      Appearance <- "[78]"
   Button "Button_79" at 263,574 size 80x46; TextOff 'EMS 79'
      on Release: ActivateScreen("711_CARRIER_STATUS", 0)
      on Press: SetTag("HMI_EMS_Nr", 79)
      ObjectEnable <- "DB16_EMS_Status_EMS_DeviceStates.DeviceStates_Condition_HMI[79]"
      Appearance <- "[79]"
   Button "Button_80" at 346,574 size 80x46; TextOff 'EMS 80'
      on Release: ActivateScreen("711_CARRIER_STATUS", 0)
      on Press: SetTag("HMI_EMS_Nr", 80)
      ObjectEnable <- "DB16_EMS_Status_EMS_DeviceStates.DeviceStates_Condition_HMI[80]"
      Appearance <- "[80]"
   Button "Button_81" at 429,574 size 80x46; TextOff 'EMS 81'
      on Release: ActivateScreen("711_CARRIER_STATUS", 0)
      on Press: SetTag("HMI_EMS_Nr", 81)
      ObjectEnable <- "DB16_EMS_Status_EMS_DeviceStates.DeviceStates_Condition_HMI[81]"
      Appearance <- "[81]"
   Button "Button_82" at 512,574 size 80x46; TextOff 'EMS 82'
      on Release: ActivateScreen("711_CARRIER_STATUS", 0)
      on Press: SetTag("HMI_EMS_Nr", 82)
      ObjectEnable <- "DB16_EMS_Status_EMS_DeviceStates.DeviceStates_Condition_HMI[82]"
      Appearance <- "[82]"
   Button "Button_83" at 595,574 size 80x46; TextOff 'Text'
   Button "Button_84" at 678,574 size 80x46; TextOff 'Text'
   Button "Button_85" at 761,574 size 80x46; TextOff 'Text'
   Button "Button_86" at 845,574 size 80x46; TextOff 'Text'
   Button "Button_87" at 928,574 size 80x46; TextOff 'Text'
   Button "Button_88" at 1011,574 size 80x46; TextOff 'Text'
   Button "Button_89" at 1094,574 size 80x46; TextOff 'Text'
   Button "Button_90" at 1178,574 size 80x46; TextOff 'Text'
   TextField "Textfeld_7" at 567,118 size 243x27; Text 'section counter / min Barcode mm / EMS Status'
   TextField "Text field_1" at 83,642 size 97x25; Text 'NO COMM'
   TextField "Text field_2" at 83,683 size 191x25; Text 'ACTIVE, NO FAULTS'
   TextField "Text field_3" at 83,722 size 90x25; Text 'FAULTED'
   TextField "Text field_4" at 83,763 size 100x25; Text 'WARNING'

screen "700_System_Line_Overview" 1280x800
   GraphicView "Graphic view_1" at 0,119 size 1144x681; Picture "LAYOUT 1"
   TextField "Text field_126" at 847,138 size 285x28; Text 'SYSTEM LAYOUT SCREEN'
   Button "Template_Button_3" at 1074,2 size 203x55; TextOn 'FAULT RESET FAULT RESET'; TextOff 'FAULT RESET FAULT RESET'
      on Release: ResetBit("DB_SDC_GLOBAL_M.SDC_ER_Reset")
      on Press: SetBit("DB_SDC_GLOBAL_M.SDC_ER_Reset")
   AlarmView "Template_Alarm view_2" at 128,2 size 948x112
   Button "Template_Button_4" at 1196,56 size 81x59; TextOff 'Text'
      Appearance <- "AlwaysTRUE"
   Button "Button_21" at 0,57 size 128x58; TextOff 'SELECT SCREEN'
      on Release: ActivateScreen("010_START", 0)
   Button "Button_22" at 0,0 size 128x58; TextOff 'PREVIOUS SCREEN'
      on Click: function_efd93a16()
   DateTimeField "Template_Date/time field_2" at 1075,56 size 123x28
   DateTimeField "Template_Date/time field_3" at 1075,83 size 122x32
   TextField "Text field_2" at 446,600 size 186x29; Text 'Line Overview 1'
   TextField "Text field_3" at 524,179 size 186x29; Text 'Line Overview 3'
   TextField "Text field_4" at 564,383 size 186x29; Text 'Line Overview 2'
   TextField "Text field_5" at 811,383 size 186x29; Text 'Line Overview 4'
   Button "Button_1" at 436,216 size 134x49; TextOn 'LINE_OVERVIEW_2 LINE OVERVIEW_2'; TextOff 'LINE_OVERVIEW_2 LINE OVERVIEW_3'
      on Click: ActivateScreen("703_Line_Overview_3", 0)
   Button "Button_2" at 592,438 size 134x49; TextOn 'LINE_OVERVIEW_2 LINE OVERVIEW_2'; TextOff 'LINE_OVERVIEW_2 LINE OVERVIEW_2'
      on Click: ActivateScreen("702_Line_Overview_2", 0)
   Button "Button_3" at 840,438 size 134x49; TextOn 'LINE_OVERVIEW_2 LINE OVERVIEW_2'; TextOff 'LINE_OVERVIEW_2 LINE OVERVIEW_4'
      on Click: ActivateScreen("704_Line_Overview_4", 0)
   Button "Button_4" at 1148,702 size 127x87; TextOn 'LINE_OVERVIEW_2 LINE OVERVIEW_2'; TextOff 'LINE_OVERVIEW_2 / Main Screen'
      on Click: ActivateScreen("010_START", 0)
   Button "Button_14" at 247,578 size 134x49; TextOn 'LINE_OVERVIEW_2 LINE OVERVIEW_2'; TextOff 'LINE_OVERVIEW_2 LINE OVERVIEW_1'
      on Click: ActivateScreen("701_Line_Overview_1", 0)

screen "LINE_OVERVIEW_1_NOT_USED" 1280x800
   GraphicView "Graphic view_1" at 79,0 size 1139x766; Picture "b1 123927_1"
   TextField "Text field_1" at 981,284 size 46x25; Text 'S14'
   TextField "Text field_2" at 901,284 size 46x25; Text 'S13'
   TextField "Text field_3" at 818,283 size 46x25; Text 'S12'
   TextField "Text field_4" at 778,283 size 46x25; Text 'S11'
   TextField "Text field_5" at 734,283 size 46x25; Text 'S10'
   TextField "Text field_6" at 696,283 size 46x25; Text 'S9'
   TextField "Text field_7" at 653,283 size 46x25; Text 'S57'
   TextField "Text field_8" at 296,283 size 46x25; Text 'S7'
   TextField "Text field_9" at 252,283 size 46x25; Text 'S6'
   TextField "Text field_10" at 154,382 size 46x25; Text 'S5'
   TextField "Text field_11" at 245,471 size 46x25; Text 'S4'
   TextField "Text field_12" at 152,437 size 46x25; Text 'S3'
   TextField "Text field_13" at 22,532 size 46x25; Text 'S2'
   TextField "Text field_14" at 13,622 size 46x25; Text 'S58'
   TextField "Text field_15" at 22,671 size 46x25; Text 'S1'
   TextField "Text field_16" at 13,707 size 46x25; Text 'S56'
   TextField "Text field_17" at 128,721 size 46x25; Text 'S55'
   TextField "Text field_18" at 249,709 size 46x25; Text 'S54'
   TextField "Text field_19" at 212,590 size 46x25; Text 'S53'
   TextField "Text field_20" at 306,590 size 46x25; Text 'S52'
   TextField "Text field_21" at 395,591 size 46x25; Text 'S51'
   TextField "Text field_22" at 473,493 size 46x25; Text 'S47'
   TextField "Text field_23" at 544,492 size 46x25; Text 'S48'
   TextField "Text field_24" at 477,674 size 46x25; Text 'S44'
   TextField "Text field_25" at 546,674 size 46x25; Text 'S43'
   TextField "Text field_26" at 622,674 size 46x25; Text 'S42'
   TextField "Text field_27" at 723,641 size 46x25; Text 'S41'
   TextField "Text field_28" at 774,523 size 46x25; Text 'S40'
   TextField "Text field_29" at 883,607 size 46x25; Text 'S39'
   TextField "Text field_30" at 1015,607 size 46x25; Text 'S38'
   TextField "Text field_31" at 1114,607 size 46x25; Text 'S37'
   TextField "Text field_32" at 1158,502 size 46x25; Text 'S36'
   TextField "Text field_33" at 1157,438 size 46x25; Text 'S35'
   TextField "Text field_34" at 1158,381 size 46x25; Text 'S34'
   TextField "Text field_35" at 33,44 size 84x24; Text 'Area Name'
   TextField "Text field_36" at 36,62 size 56x25; Text 'Area A'
   Button "Button_14" at 980,678 size 140x105; TextOn 'LINE_OVERVIEW_2 LINE OVERVIEW_2'; TextOff 'LINE_OVERVIEW_2 LINE OVERVIEW_2'
      on Click: ActivateScreen("LINE_OVERVIEW_2_NOT_USED", 0)
   Button "Button_1" at 1125,677 size 140x105; TextOn 'LINE_OVERVIEW_2 LINE OVERVIEW_2'; TextOff 'LINE_OVERVIEW_2 / Main Screen'
      on Click: ActivateScreen("010_START", 0)
   TextField "Text field_37" at 36,78 size 67x25; Text 'Area AA'
   TextField "Text field_38" at 36,94 size 55x25; Text 'Area B'
   TextField "Text field_39" at 36,112 size 65x25; Text 'Area BB'
   TextField "Text field_40" at 36,129 size 55x25; Text 'Area C'
   TextField "Text field_41" at 36,147 size 65x25; Text 'Area CC'
   TextField "Text field_42" at 36,165 size 56x25; Text 'Area H'
   TextField "Text field_43" at 36,182 size 57x25; Text 'Area D'
   TextField "Text field_44" at 36,200 size 55x25; Text 'Area E'
   TextField "Text field_45" at 36,218 size 54x25; Text 'Area F'
   TextField "Text field_46" at 36,237 size 63x25; Text 'Area FF'
   TextField "Text field_47" at 36,256 size 56x25; Text 'Area G'
   TextField "Text field_48" at 242,42 size 81x26; Text 'Area Start'
   TextField "Text field_49" at 241,61 size 109x25; Text 'After Cab Pick'
   TextField "Text field_50" at 241,77 size 39x25; Text 'DL 1'
   TextField "Text field_51" at 241,94 size 155x25; Text 'DL 2 (Marriege Cell)'
   TextField "Text field_52" at 240,111 size 166x25; Text 'S14 at 90 degree turn'
   TextField "Text field_53" at 240,128 size 123x25; Text 'S16 Check Point'
   TextField "Text field_54" at 240,147 size 187x25; Text 'S19 above Front Bumper'
   TextField "Text field_55" at 240,164 size 125x25; Text 'from the Shuttle'
   TextField "Text field_56" at 240,181 size 169x25; Text 'S32 at 90 Degree turn'
   TextField "Text field_57" at 240,200 size 192x25; Text 'S33 at EMS01 Main Panel'
   TextField "Text field_58" at 240,219 size 198x25; Text 'S36 before 90 degree turn'
   TextField "Text field_59" at 241,237 size 106x25; Text 'Before Repair'
   TextField "Text field_60" at 241,255 size 91x25; Text 'Repair Spur'
   TextField "Text field_61" at 445,43 size 73x26; Text 'Area End'
   TextField "Text field_62" at 445,62 size 38x25; Text 'DL1'
   TextField "Text field_63" at 445,77 size 155x25; Text 'DL 2 (Marriege Cell)'
   TextField "Text field_64" at 445,95 size 166x25; Text 'S14 at 90 degree turn'
   TextField "Text field_65" at 445,113 size 123x25; Text 'S16 Check Point'
   TextField "Text field_66" at 445,130 size 187x25; Text 'S19 above Front Bumper'
   TextField "Text field_67" at 445,147 size 139x25; Text 'Before the Shuttle'
   TextField "Text field_68" at 444,165 size 169x25; Text 'S32 at 90 Degree turn'
   TextField "Text field_69" at 444,183 size 192x25; Text 'S33 at EMS01 Main Panel'
   TextField "Text field_70" at 444,201 size 198x25; Text 'S36 before 90 degree turn'
   TextField "Text field_71" at 445,220 size 106x25; Text 'Before Repair'
   TextField "Text field_72" at 446,238 size 67x25; Text 'Cab Pick'
   TextField "Text field_73" at 446,255 size 91x25; Text 'Repair Spur'
   TextField "Text field_74" at 652,43 size 67x26; Text 'Location'
   TextField "Text field_75" at 651,62 size 45x25; Text '@G7'
   TextField "Text field_76" at 651,79 size 47x25; Text '@F14'
   TextField "Text field_77" at 651,96 size 47x25; Text '@F14'
   TextField "Text field_78" at 651,112 size 50x25; Text '@Q16'
   TextField "Text field_79" at 651,131 size 50x25; Text '@Q16'
   TextField "Text field_80" at 651,149 size 49x25; Text '@U12'
   TextField "Text field_81" at 651,167 size 49x25; Text '@U12'
   TextField "Text field_82" at 651,184 size 46x25; Text '@L17'
   TextField "Text field_83" at 651,202 size 46x25; Text '@L17'
   TextField "Text field_84" at 651,221 size 48x25; Text '@C17'
   TextField "Text field_85" at 651,239 size 41x25; Text '@D9'
   TextField "Text field_86" at 651,257 size 41x25; Text '@D9'
   TextField "Text field_87" at 737,42 size 45x26; Text 'Panel'
   TextField "Text field_88" at 736,62 size 115x25; Text 'EMS01R2 JB33'
   TextField "Text field_89" at 736,80 size 75x25; Text 'EMS01R3'
   TextField "Text field_90" at 736,97 size 75x25; Text 'EMS01R3'
   TextField "Text field_91" at 736,113 size 100x25; Text 'EMS01 JB22'
   TextField "Text field_92" at 736,130 size 95x25; Text 'EMS01 JB22'
   TextField "Text field_93" at 736,148 size 75x25; Text 'EMS01R4'
   TextField "Text field_94" at 736,167 size 75x25; Text 'EMS01R4'
   TextField "Text field_95" at 736,185 size 55x25; Text 'EMS01'
   TextField "Text field_96" at 737,202 size 55x25; Text 'EMS01'
   TextField "Text field_97" at 737,220 size 115x25; Text 'EMS01R1 JB23'
   TextField "Text field_98" at 737,238 size 75x25; Text 'EMS01R1'
   TextField "Text field_99" at 737,256 size 75x25; Text 'EMS01R1'
   TextField "Text field_100" at 906,43 size 50x26; Text 'Offset'
   TextField "Text field_101" at 907,62 size 38x25; Text '9'
   TextField "Text field_102" at 907,80 size 38x25; Text '1'
   TextField "Text field_103" at 907,98 size 38x25; Text '2'
   TextField "Text field_104" at 907,114 size 38x25; Text '10'
   TextField "Text field_105" at 907,130 size 38x25; Text '11'
   TextField "Text field_106" at 907,150 size 38x25; Text '3'
   TextField "Text field_107" at 907,168 size 38x25; Text '4'
   TextField "Text field_108" at 907,185 size 38x25; Text '5'
   TextField "Text field_109" at 907,202 size 38x25; Text '6'
   TextField "Text field_110" at 907,221 size 38x25; Text '7'
   TextField "Text field_111" at 908,238 size 38x25; Text '12'
   TextField "Text field_112" at 908,256 size 38x25; Text '8'
   TextField "Text field_113" at 1084,54 size 82x22; Text 'AREA BB'
   TextField "Text field_114" at 1131,251 size 71x22; Text 'AREA E'
   TextField "Text field_115" at 940,613 size 71x22; Text 'AREA F'
   TextField "Text field_116" at 493,464 size 71x22; Text 'AREA G'
   TextField "Text field_117" at 267,679 size 82x22; Text 'AREA FF'
   TextField "Text field_118" at 138,519 size 71x22; Text 'AREA A'
   TextField "Text field_119" at 515,360 size 82x22; Text 'AREA AA'
   TextField "Text field_120" at 950,362 size 71x22; Text 'AREA B'
   TextField "Text field_121" at 731,358 size 53x27; Text 'DL2'
   TextField "Text field_122" at 712,381 size 93x25; Text 'Mrg Cell'
   TextField "Text field_123" at 296,359 size 53x27; Text 'DL1'
   TextField "Text field_124" at 125,635 size 49x25; Text 'Cab'
   TextField "Text field_125" at 125,656 size 49x25; Text 'Pick'
   TextField "Text field_126" at 454,13 size 341x28; Text 'OVERVIEW 1 - SCREEN 0023'
   TextField "Text field_127" at 614,387 size 82x24; Text 'EMS01R3'
   TextField "Text field_128" at 614,421 size 82x22; Text 'AREA AA'
   TextField "Text field_129" at 619,452 size 71x22; Text 'AREA B'
   TextField "Text field_130" at 23,313 size 82x24; Text 'EMS01R2'
   TextField "Text field_131" at 38,329 size 49x24; Text 'JB33'
   TextField "Text field_132" at 28,361 size 71x22; Text 'AREA A'
   TextField "Text field_133" at 379,679 size 82x24; Text 'EMS01R1'
   TextField "Text field_134" at 385,702 size 71x22; Text 'AREA G'
   TextField "Text field_135" at 386,729 size 71x22; Text 'AREA F'
   TextField "Text field_136" at 380,754 size 82x22; Text 'AREA FF'
   TextField "Text field_137" at 703,687 size 60x24; Text 'EMS01'
   TextField "Text field_138" at 699,718 size 71x22; Text 'AREA D'
   TextField "Text field_139" at 699,746 size 71x22; Text 'AREA E'
   TextField "Text field_140" at 790,686 size 82x24; Text 'EMS01R4'
   TextField "Text field_143" at 897,679 size 60x24; Text 'EMS01'
   TextField "Text field_144" at 902,693 size 49x24; Text 'JB22'
   DateTimeField "Date/time field_1" at 11,12 size 258x34
   TextField "Text field_141" at 790,718 size 82x22; Text 'AREA CC'
   TextField "Text field_142" at 796,746 size 71x22; Text 'AREA H'
   TextField "Text field_146" at 891,745 size 71x22; Text 'AREA C'
   TextField "Text field_145" at 886,718 size 82x22; Text 'AREA BB'
   TextField "Text field_147" at 863,43 size 38x26; Text 'Slot'
   TextField "Text field_148" at 865,62 size 38x25; Text '13'
   TextField "Text field_149" at 865,80 size 38x25; Text '5'
   TextField "Text field_150" at 865,97 size 38x25; Text '6'
   TextField "Text field_151" at 865,113 size 38x25; Text '14'
   TextField "Text field_152" at 865,131 size 38x25; Text '15'
   TextField "Text field_153" at 865,150 size 38x25; Text '7'
   TextField "Text field_154" at 865,166 size 38x25; Text '12'
   TextField "Text field_155" at 865,184 size 38x25; Text '8'
   TextField "Text field_156" at 865,202 size 38x25; Text '9'
   TextField "Text field_157" at 865,220 size 38x25; Text '10'
   TextField "Text field_158" at 866,238 size 38x25; Text '16'
   TextField "Text field_159" at 866,256 size 38x25; Text '11'
   TextField "Text field_160" at 120,43 size 40x26; Text 'Area'
   TextField "Text field_161" at 118,62 size 98x25; Text 'Cab Delivery'
   TextField "Text field_162" at 118,78 size 53x25; Text 'Trim 5'
   TextField "Text field_163" at 118,93 size 106x25; Text 'Body Delivery'
   TextField "Text field_164" at 118,110 size 106x25; Text 'Body Delivery'
   TextField "Text field_165" at 118,127 size 106x25; Text 'Body Delivery'
   TextField "Text field_166" at 118,146 size 106x25; Text 'Body Delivery'
   TextField "Text field_167" at 118,164 size 83x25; Text 'Body Deck'
   TextField "Text field_168" at 118,181 size 107x25; Text 'Empty Return'
   TextField "Text field_169" at 118,200 size 107x25; Text 'Empty Return'
   TextField "Text field_170" at 118,218 size 107x25; Text 'Empty Return'
   TextField "Text field_171" at 118,236 size 107x25; Text 'Empty Return'
   TextField "Text field_172" at 116,255 size 91x25; Text 'Repair Spur'
   IOField "I/O field_42" at 129,761 size 37x32; FormatPattern 99
      ProcessValue <- "CarrierNumber"
   IOField "I/O field_1" at 56,703 size 37x32; FormatPattern 99
      ProcessValue <- "CarrierNumber"
   IOField "I/O field_2" at 56,666 size 37x32; FormatPattern 99
      ProcessValue <- "CarrierNumber"
   IOField "I/O field_3" at 56,617 size 37x32; FormatPattern 99
      ProcessValue <- "CarrierNumber"
   IOField "I/O field_4" at 56,568 size 37x32; FormatPattern 99
      ProcessValue <- "CarrierNumber"
   IOField "I/O field_5" at 56,527 size 37x32; FormatPattern 99
      ProcessValue <- "CarrierNumber"
   IOField "I/O field_6" at 106,467 size 37x32; FormatPattern 99
      ProcessValue <- "CarrierNumber"
   IOField "I/O field_7" at 148,467 size 37x32; FormatPattern 99
      ProcessValue <- "CarrierNumber"
   IOField "I/O field_8" at 190,467 size 37x32; FormatPattern 99
      ProcessValue <- "CarrierNumber"
   IOField "I/O field_9" at 191,413 size 37x32; FormatPattern 99
      ProcessValue <- "CarrierNumber"
   IOField "I/O field_10" at 191,378 size 37x32; FormatPattern 99
      ProcessValue <- "CarrierNumber"
   IOField "I/O field_11" at 248,310 size 37x32; FormatPattern 99
      ProcessValue <- "CarrierNumber"
   IOField "I/O field_12" at 292,310 size 37x32; FormatPattern 99
      ProcessValue <- "CarrierNumber"
   IOField "I/O field_13" at 337,310 size 37x32; FormatPattern 99
      ProcessValue <- "CarrierNumber"
   IOField "I/O field_14" at 376,310 size 37x32; FormatPattern 99
      ProcessValue <- "CarrierNumber"
   IOField "I/O field_15" at 415,310 size 37x32; FormatPattern 99
      ProcessValue <- "CarrierNumber"
   IOField "I/O field_16" at 453,310 size 37x32; FormatPattern 99
      ProcessValue <- "CarrierNumber"
   IOField "I/O field_17" at 492,310 size 37x32; FormatPattern 99
      ProcessValue <- "CarrierNumber"
   IOField "I/O field_18" at 531,310 size 37x32; FormatPattern 99
      ProcessValue <- "CarrierNumber"
   IOField "I/O field_19" at 570,310 size 37x32; FormatPattern 99
      ProcessValue <- "CarrierNumber"
   IOField "I/O field_20" at 609,310 size 37x32; FormatPattern 99
      ProcessValue <- "CarrierNumber"
   IOField "I/O field_21" at 654,310 size 37x32; FormatPattern 99
      ProcessValue <- "CarrierNumber"
   IOField "I/O field_22" at 692,310 size 37x32; FormatPattern 99
      ProcessValue <- "CarrierNumber"
   IOField "I/O field_23" at 736,310 size 37x32; FormatPattern 99
      ProcessValue <- "CarrierNumber"
   IOField "I/O field_24" at 778,310 size 37x32; FormatPattern 99
      ProcessValue <- "CarrierNumber"
   IOField "I/O field_25" at 819,310 size 37x32; FormatPattern 99
      ProcessValue <- "CarrierNumber"
   IOField "I/O field_26" at 863,310 size 37x32; FormatPattern 99
      ProcessValue <- "CarrierNumber"
   IOField "I/O field_27" at 902,310 size 37x32; FormatPattern 99
      ProcessValue <- "CarrierNumber"
   IOField "I/O field_28" at 945,310 size 37x32; FormatPattern 99
      ProcessValue <- "CarrierNumber"
   IOField "I/O field_29" at 984,310 size 37x32; FormatPattern 99
      ProcessValue <- "CarrierNumber"
   IOField "I/O field_30" at 1031,289 size 37x32; FormatPattern 99
      ProcessValue <- "CarrierNumber"
   IOField "I/O field_31" at 1031,257 size 37x32; FormatPattern 99
      ProcessValue <- "CarrierNumber"
   IOField "I/O field_32" at 1031,225 size 37x32; FormatPattern 99
      ProcessValue <- "CarrierNumber"
   IOField "I/O field_33" at 1031,193 size 37x32; FormatPattern 99
      ProcessValue <- "CarrierNumber"
   IOField "I/O field_34" at 1031,162 size 37x32; FormatPattern 99
      ProcessValue <- "CarrierNumber"
   IOField "I/O field_35" at 1031,131 size 37x32; FormatPattern 99
      ProcessValue <- "CarrierNumber"
   IOField "I/O field_36" at 1031,99 size 37x32; FormatPattern 99
      ProcessValue <- "CarrierNumber"
   IOField "I/O field_37" at 1031,67 size 37x32; FormatPattern 99
      ProcessValue <- "CarrierNumber"
   IOField "I/O field_38" at 1031,35 size 37x32; FormatPattern 99
      ProcessValue <- "CarrierNumber"
   IOField "I/O field_39" at 1031,3 size 37x32; FormatPattern 99
      ProcessValue <- "CarrierNumber"
   IOField "I/O field_49" at 1219,339 size 37x32; FormatPattern 99
      ProcessValue <- "CarrierNumber"
   IOField "I/O field_50" at 1219,378 size 37x32; FormatPattern 99
      ProcessValue <- "CarrierNumber"
   IOField "I/O field_51" at 1219,435 size 37x32; FormatPattern 99
      ProcessValue <- "CarrierNumber"
   IOField "I/O field_52" at 1218,498 size 37x32; FormatPattern 99
      ProcessValue <- "CarrierNumber"
   IOField "I/O field_40" at 1218,302 size 37x32; FormatPattern 99
      ProcessValue <- "CarrierNumber"
   IOField "I/O field_41" at 1218,265 size 37x32; FormatPattern 99
      ProcessValue <- "CarrierNumber"
   IOField "I/O field_43" at 1218,228 size 37x32; FormatPattern 99
      ProcessValue <- "CarrierNumber"
   IOField "I/O field_44" at 1218,191 size 37x32; FormatPattern 99
      ProcessValue <- "CarrierNumber"
   IOField "I/O field_45" at 1218,154 size 37x32; FormatPattern 99
      ProcessValue <- "CarrierNumber"
   IOField "I/O field_46" at 1218,117 size 37x32; FormatPattern 99
      ProcessValue <- "CarrierNumber"
   IOField "I/O field_47" at 1218,80 size 37x32; FormatPattern 99
      ProcessValue <- "CarrierNumber"
   IOField "I/O field_48" at 1218,43 size 37x32; FormatPattern 99
      ProcessValue <- "CarrierNumber"
   IOField "I/O field_53" at 1156,568 size 37x32; FormatPattern 99
      ProcessValue <- "CarrierNumber"
   IOField "I/O field_54" at 1115,568 size 37x32; FormatPattern 99
      ProcessValue <- "CarrierNumber"
   IOField "I/O field_55" at 1054,568 size 37x32; FormatPattern 99
      ProcessValue <- "CarrierNumber"
   IOField "I/O field_56" at 1015,568 size 37x32; FormatPattern 99
      ProcessValue <- "CarrierNumber"
   IOField "I/O field_57" at 924,568 size 37x32; FormatPattern 99
      ProcessValue <- "CarrierNumber"
   IOField "I/O field_58" at 884,568 size 37x32; FormatPattern 99
      ProcessValue <- "CarrierNumber"
   IOField "I/O field_59" at 813,568 size 37x32; FormatPattern 99
      ProcessValue <- "CarrierNumber"
   IOField "I/O field_60" at 773,568 size 37x32; FormatPattern 99
      ProcessValue <- "CarrierNumber"
   IOField "I/O field_61" at 724,603 size 37x32; FormatPattern 99
      ProcessValue <- "CarrierNumber"
   IOField "I/O field_62" at 663,634 size 37x32; FormatPattern 99
      ProcessValue <- "CarrierNumber"
   IOField "I/O field_63" at 622,634 size 37x32; FormatPattern 99
      ProcessValue <- "CarrierNumber"
   IOField "I/O field_64" at 545,527 size 37x32; FormatPattern 99
      ProcessValue <- "CarrierNumber"
   IOField "I/O field_65" at 475,527 size 37x32; FormatPattern 99
      ProcessValue <- "CarrierNumber"
   IOField "I/O field_66" at 548,632 size 37x32; FormatPattern 99
      ProcessValue <- "CarrierNumber"
   IOField "I/O field_67" at 478,632 size 37x32; FormatPattern 99
      ProcessValue <- "CarrierNumber"
   IOField "I/O field_68" at 399,632 size 37x32; FormatPattern 99
      ProcessValue <- "CarrierNumber"
   IOField "I/O field_69" at 348,632 size 37x32; FormatPattern 99
      ProcessValue <- "CarrierNumber"
   IOField "I/O field_70" at 306,632 size 37x32; FormatPattern 99
      ProcessValue <- "CarrierNumber"
   IOField "I/O field_71" at 255,632 size 37x32; FormatPattern 99
      ProcessValue <- "CarrierNumber"
   IOField "I/O field_72" at 214,632 size 37x32; FormatPattern 99
      ProcessValue <- "CarrierNumber"
   IOField "I/O field_73" at 202,671 size 37x32; FormatPattern 99
      ProcessValue <- "CarrierNumber"
   IOField "I/O field_74" at 202,707 size 37x32; FormatPattern 99
      ProcessValue <- "CarrierNumber"

screen "LINE_OVERVIEW_2_NOT_USED" 1280x800
   IOField "I/O field_1" at 299,73 size 37x32; FormatPattern 99
      ProcessValue <- "CarrierNumber"
   IOField "I/O field_2" at 186,73 size 37x32; FormatPattern 99
      ProcessValue <- "CarrierNumber"
   IOField "I/O field_3" at 54,139 size 37x32; FormatPattern 99
      ProcessValue <- "CarrierNumber"
   IOField "I/O field_4" at 232,73 size 37x32; FormatPattern 99
      ProcessValue <- "CarrierNumber"
   IOField "I/O field_5" at 299,36 size 37x32; FormatPattern 99
      ProcessValue <- "CarrierNumber"
   IOField "I/O field_6" at 142,73 size 37x32; FormatPattern 99
      ProcessValue <- "CarrierNumber"
   IOField "I/O field_7" at 362,73 size 37x32; FormatPattern 99
      ProcessValue <- "CarrierNumber"
   IOField "I/O field_8" at 435,73 size 37x32; FormatPattern 99
      ProcessValue <- "CarrierNumber"
   IOField "I/O field_9" at 512,73 size 37x32; FormatPattern 99
      ProcessValue <- "CarrierNumber"
   IOField "I/O field_10" at 598,73 size 37x32; FormatPattern 99
      ProcessValue <- "CarrierNumber"
   IOField "I/O field_11" at 685,73 size 37x32; FormatPattern 99
      ProcessValue <- "CarrierNumber"
   IOField "I/O field_12" at 782,73 size 37x32; FormatPattern 99
      ProcessValue <- "CarrierNumber"
   IOField "I/O field_13" at 836,73 size 37x32; FormatPattern 99
      ProcessValue <- "CarrierNumber"
   IOField "I/O field_14" at 934,73 size 37x32; FormatPattern 99
      ProcessValue <- "CarrierNumber"
   IOField "I/O field_15" at 992,73 size 37x32; FormatPattern 99
      ProcessValue <- "CarrierNumber"
   IOField "I/O field_16" at 1086,104 size 37x32; FormatPattern 99
      ProcessValue <- "CarrierNumber"
   IOField "I/O field_17" at 1086,137 size 37x32; FormatPattern 99
      ProcessValue <- "CarrierNumber"
   IOField "I/O field_18" at 1086,170 size 37x32; FormatPattern 99
      ProcessValue <- "CarrierNumber"
   IOField "I/O field_19" at 1086,203 size 37x32; FormatPattern 99
      ProcessValue <- "CarrierNumber"
   IOField "I/O field_20" at 1086,236 size 37x32; FormatPattern 99
      ProcessValue <- "CarrierNumber"
   IOField "I/O field_21" at 1086,269 size 37x32; FormatPattern 99
      ProcessValue <- "CarrierNumber"
   IOField "I/O field_22" at 1086,302 size 37x32; FormatPattern 99
      ProcessValue <- "CarrierNumber"
   IOField "I/O field_23" at 1086,335 size 37x32; FormatPattern 99
      ProcessValue <- "CarrierNumber"
   IOField "I/O field_24" at 1086,368 size 37x32; FormatPattern 99
      ProcessValue <- "CarrierNumber"
   IOField "I/O field_25" at 1086,401 size 37x32; FormatPattern 99
      ProcessValue <- "CarrierNumber"
   IOField "I/O field_26" at 1086,434 size 37x32; FormatPattern 99
      ProcessValue <- "CarrierNumber"
   IOField "I/O field_27" at 1086,467 size 37x32; FormatPattern 99
      ProcessValue <- "CarrierNumber"
   IOField "I/O field_28" at 1086,500 size 37x32; FormatPattern 99
      ProcessValue <- "CarrierNumber"
   IOField "I/O field_29" at 1086,533 size 37x32; FormatPattern 99
      ProcessValue <- "CarrierNumber"
   IOField "I/O field_30" at 1086,566 size 37x32; FormatPattern 99
      ProcessValue <- "CarrierNumber"
   IOField "I/O field_31" at 1086,599 size 37x32; FormatPattern 99
      ProcessValue <- "CarrierNumber"
   IOField "I/O field_32" at 1086,637 size 37x32; FormatPattern 99
      ProcessValue <- "CarrierNumber"
   IOField "I/O field_33" at 1086,669 size 37x32; FormatPattern 99
      ProcessValue <- "CarrierNumber"
   IOField "I/O field_34" at 1086,701 size 37x32; FormatPattern 99
      ProcessValue <- "CarrierNumber"
   IOField "I/O field_35" at 1086,733 size 37x32; FormatPattern 99
      ProcessValue <- "CarrierNumber"
   IOField "I/O field_36" at 1086,765 size 37x32; FormatPattern 99
      ProcessValue <- "CarrierNumber"
   IOField "I/O field_37" at 142,207 size 37x32; FormatPattern 99
      ProcessValue <- "CarrierNumber"
   IOField "I/O field_38" at 186,208 size 37x32; FormatPattern 99
      ProcessValue <- "CarrierNumber"
   IOField "I/O field_39" at 230,208 size 37x32; FormatPattern 99
      ProcessValue <- "CarrierNumber"
   IOField "I/O field_40" at 274,208 size 37x32; FormatPattern 99
      ProcessValue <- "CarrierNumber"
   IOField "I/O field_41" at 318,208 size 37x32; FormatPattern 99
      ProcessValue <- "CarrierNumber"
   IOField "I/O field_42" at 362,208 size 37x32; FormatPattern 99
      ProcessValue <- "CarrierNumber"
   IOField "I/O field_43" at 406,208 size 37x32; FormatPattern 99
      ProcessValue <- "CarrierNumber"
   IOField "I/O field_44" at 450,208 size 37x32; FormatPattern 99
      ProcessValue <- "CarrierNumber"
   IOField "I/O field_45" at 544,208 size 37x32; FormatPattern 99
      ProcessValue <- "CarrierNumber"
   IOField "I/O field_46" at 592,208 size 37x32; FormatPattern 99
      ProcessValue <- "CarrierNumber"
   IOField "I/O field_47" at 684,207 size 37x32; FormatPattern 99
      ProcessValue <- "CarrierNumber"
   IOField "I/O field_48" at 730,207 size 37x32; FormatPattern 99
      ProcessValue <- "CarrierNumber"
   IOField "I/O field_49" at 803,236 size 37x32; FormatPattern 99
      ProcessValue <- "CarrierNumber"
   IOField "I/O field_50" at 803,268 size 37x32; FormatPattern 99
      ProcessValue <- "CarrierNumber"
   IOField "I/O field_51" at 803,300 size 37x32; FormatPattern 99
      ProcessValue <- "CarrierNumber"
   IOField "I/O field_52" at 803,332 size 37x32; FormatPattern 99
      ProcessValue <- "CarrierNumber"
   IOField "I/O field_53" at 803,364 size 37x32; FormatPattern 99
      ProcessValue <- "CarrierNumber"
   IOField "I/O field_54" at 803,396 size 37x32; FormatPattern 99
      ProcessValue <- "CarrierNumber"
   IOField "I/O field_55" at 803,436 size 37x32; FormatPattern 99
      ProcessValue <- "CarrierNumber"
   IOField "I/O field_56" at 803,475 size 37x32; FormatPattern 99
      ProcessValue <- "CarrierNumber"
   IOField "I/O field_57" at 803,507 size 37x32; FormatPattern 99
      ProcessValue <- "CarrierNumber"
   IOField "I/O field_58" at 803,539 size 37x32; FormatPattern 99
      ProcessValue <- "CarrierNumber"
   IOField "I/O field_59" at 803,571 size 37x32; FormatPattern 99
      ProcessValue <- "CarrierNumber"
   IOField "I/O field_60" at 803,603 size 37x32; FormatPattern 99
      ProcessValue <- "CarrierNumber"
   IOField "I/O field_61" at 803,635 size 37x32; FormatPattern 99
      ProcessValue <- "CarrierNumber"
   IOField "I/O field_62" at 803,667 size 37x32; FormatPattern 99
      ProcessValue <- "CarrierNumber"
   IOField "I/O field_63" at 803,699 size 37x32; FormatPattern 99
      ProcessValue <- "CarrierNumber"
   IOField "I/O field_64" at 803,731 size 37x32; FormatPattern 99
      ProcessValue <- "CarrierNumber"
   IOField "I/O field_65" at 803,763 size 37x32; FormatPattern 99
      ProcessValue <- "CarrierNumber"
   GraphicView "Graphic view_1" at 67,88 size 1015x709; Picture "b2 124337_2"
   TextField "Text field_1" at 858,242 size 46x25; Text 'S17'
   TextField "Text field_2" at 858,441 size 46x25; Text 'S16'
   TextField "Text field_3" at 858,479 size 46x25; Text 'S15'
   TextField "Text field_4" at 1028,604 size 46x25; Text 'S33'
   TextField "Text field_5" at 989,40 size 46x25; Text 'S32'
   TextField "Text field_6" at 833,40 size 46x25; Text 'S31'
   TextField "Text field_7" at 683,40 size 46x25; Text 'S30'
   TextField "Text field_8" at 597,40 size 46x25; Text 'S29'
   TextField "Text field_9" at 511,40 size 46x25; Text 'S28'
   TextField "Text field_10" at 434,40 size 46x25; Text 'S27'
   TextField "Text field_11" at 359,40 size 46x25; Text 'S26'
   TextField "Text field_12" at 297,6 size 46x25; Text 'S24'
   TextField "Text field_13" at 296,119 size 46x25; Text 'S23'
   TextField "Text field_14" at 231,41 size 46x25; Text 'S22'
   TextField "Text field_15" at 8,141 size 46x25; Text 'S21'
   TextField "Text field_16" at 140,247 size 46x25; Text 'S20'
   TextField "Text field_17" at 543,245 size 46x25; Text 'S19'
   TextField "Text field_18" at 683,244 size 46x25; Text 'S18'
   Button "Button_14" at 1140,106 size 127x84; TextOn 'LINE_OVERVIEW_2 LINE OVERVIEW_2'; TextOff 'LINE_OVERVIEW_2 LINE OVERVIEW_1'
      on Click: ActivateScreen("LINE_OVERVIEW_1_NOT_USED", 0)
   Button "Button_1" at 1140,13 size 127x87; TextOn 'LINE_OVERVIEW_2 LINE OVERVIEW_2'; TextOff 'LINE_OVERVIEW_2 / Main Screen'
      on Click: ActivateScreen("010_START", 0)
   TextField "Text field_36" at 25,413 size 45x26; Text 'Area'
   TextField "Text field_19" at 23,431 size 56x25; Text 'Area A'
   TextField "Text field_20" at 23,446 size 67x25; Text 'Area AA'
   TextField "Text field_21" at 23,461 size 55x25; Text 'Area B'
   TextField "Text field_22" at 23,477 size 65x25; Text 'Area BB'
   TextField "Text field_23" at 23,493 size 55x25; Text 'Area C'
   TextField "Text field_24" at 23,510 size 65x25; Text 'Area CC'
   TextField "Text field_25" at 23,527 size 56x25; Text 'Area H'
   TextField "Text field_26" at 23,543 size 57x25; Text 'Area D'
   TextField "Text field_27" at 23,559 size 55x25; Text 'Area E'
   TextField "Text field_28" at 23,575 size 54x25; Text 'Area F'
   TextField "Text field_29" at 23,591 size 63x25; Text 'Area FF'
   TextField "Text field_30" at 23,609 size 56x25; Text 'Area G'
   TextField "Text field_31" at 115,413 size 88x26; Text 'Area Name'
   TextField "Text field_32" at 114,432 size 98x25; Text 'Cab Delivery'
   TextField "Text field_33" at 114,446 size 53x25; Text 'Trim 5'
   TextField "Text field_40" at 114,527 size 83x25; Text 'Body Deck'
   TextField "Text field_41" at 114,542 size 107x25; Text 'Empty Return'
   TextField "Text field_42" at 114,558 size 107x25; Text 'Empty Return'
   TextField "Text field_43" at 114,574 size 107x25; Text 'Empty Return'
   TextField "Text field_44" at 114,590 size 107x25; Text 'Empty Return'
   TextField "Text field_51" at 244,526 size 125x25; Text 'from the Shuttle'
   TextField "Text field_53" at 244,557 size 192x25; Text 'S33 at EMS01 Main Panel'
   TextField "Text field_55" at 244,591 size 106x25; Text 'Before Repair'
   TextField "Text field_56" at 244,608 size 91x25; Text 'Repair Spur'
   TextField "Text field_58" at 456,415 size 73x26; Text 'Area End'
   TextField "Text field_59" at 457,434 size 39x25; Text 'DL 1'
   TextField "Text field_60" at 457,448 size 155x25; Text 'DL 2 (Marriege Cell)'
   TextField "Text field_61" at 456,463 size 173x25; Text 'S14 at 90 Degree Turn'
   TextField "Text field_62" at 456,479 size 123x25; Text 'S16 Check Point'
   TextField "Text field_63" at 456,495 size 189x25; Text 'S19 Above Front Bumper'
   TextField "Text field_64" at 457,511 size 139x25; Text 'Before the Shuttle'
   TextField "Text field_65" at 456,526 size 173x25; Text 'S32 at 90 Degree Turn'
   TextField "Text field_66" at 456,542 size 192x25; Text 'S33 at EMS01 Main Panel'
   TextField "Text field_67" at 456,558 size 206x25; Text 'S36 Before 90 Degree Turn'
   TextField "Text field_68" at 457,575 size 106x25; Text 'Before Repair'
   TextField "Text field_69" at 457,592 size 67x25; Text 'Cab Pick'
   TextField "Text field_70" at 457,608 size 91x25; Text 'Repair Spur'
   TextField "Text field_126" at 505,4 size 341x28; Text 'OVERVIEW 2 - SCREEN 0024'
   TextField "Text field_117" at 1143,770 size 71x22; Text 'AREA E'
   TextField "Text field_71" at 1146,391 size 71x22; Text 'AREA D'
   TextField "Text field_72" at 838,132 size 71x22; Text 'AREA H'
   TextField "Text field_73" at 119,144 size 82x22; Text 'AREA CC'
   TextField "Text field_74" at 711,287 size 71x24; Text 'AREA C'
   TextField "Text field_75" at 867,706 size 82x22; Text 'AREA BB'
   TextField "Text field_121" at 504,129 size 61x28; Text 'DL5'
   TextField "Text field_76" at 512,308 size 82x24; Text 'EMS01R4'
   TextField "Text field_77" at 511,337 size 82x22; Text 'AREA CC'
   TextField "Text field_78" at 516,365 size 71x22; Text 'AREA H'
   TextField "Text field_79" at 943,303 size 60x24; Text 'EMS01'
   TextField "Text field_80" at 946,317 size 49x24; Text 'JB22'
   TextField "Text field_81" at 930,344 size 82x22; Text 'AREA BB'
   TextField "Text field_82" at 935,375 size 71x22; Text 'AREA C'
   TextField "Text field_83" at 14,647 size 82x24; Text 'EMS01R2'
   TextField "Text field_84" at 28,663 size 49x24; Text 'JB33'
   TextField "Text field_85" at 20,691 size 71x22; Text 'AREA A'
   TextField "Text field_86" at 107,644 size 82x24; Text 'EMS01R1'
   TextField "Text field_87" at 112,664 size 71x22; Text 'AREA G'
   TextField "Text field_88" at 112,690 size 71x22; Text 'AREA F'
   TextField "Text field_89" at 107,717 size 82x22; Text 'AREA FF'
   TextField "Text field_90" at 203,648 size 82x24; Text 'EMS01R3'
   TextField "Text field_91" at 203,678 size 82x22; Text 'AREA AA'
   TextField "Text field_92" at 208,711 size 71x22; Text 'AREA B'
   TextField "Text field_93" at 1161,577 size 60x24; Text 'EMS01'
   TextField "Text field_94" at 1156,610 size 71x22; Text 'AREA D'
   TextField "Text field_95" at 1155,638 size 71x22; Text 'AREA E'
   TextField "Text field_96" at 362,5 size 131x28; Text 'Body Deck'
   TextField "Text field_39" at 115,607 size 91x25; Text 'Repair Spur'
   DateTimeField "Date/time field_1" at 12,5 size 258x34
   TextField "Text field_54" at 244,575 size 206x25; Text 'S36 Before 90 Degree Turn'
   TextField "Text field_38" at 114,511 size 106x25; Text 'Body Delivery'
   TextField "Text field_37" at 114,494 size 106x25; Text 'Body Delivery'
   TextField "Text field_35" at 114,477 size 106x25; Text 'Body Delivery'
   TextField "Text field_34" at 114,462 size 106x25; Text 'Body Delivery'
   TextField "Text field_45" at 244,414 size 81x26; Text 'Area Start'
   TextField "Text field_46" at 244,431 size 109x25; Text 'After Cab Pick'
   TextField "Text field_47" at 244,445 size 39x25; Text 'DL 1'
   TextField "Text field_48" at 244,461 size 155x25; Text 'DL 2 (Marriege Cell)'
   TextField "Text field_49" at 244,477 size 173x25; Text 'S14 at 90 Degree Turn'
   TextField "Text field_50" at 244,494 size 123x25; Text 'S16 Check Point'
   TextField "Text field_52" at 244,542 size 173x25; Text 'S32 at 90 Degree Turn'
   TextField "Text field_57" at 244,511 size 189x25; Text 'S19 Above Front Bumper'

screen "707_GLOBAL_PARAMETER" 1280x800, template "Top_Header"
   on GenerateScreen: SetTag("SDC\_intern_Bildnummer", 700)
   IOField "EA-Feld_10" at 373,350 size 122x32; FormatPattern 99999999
      Appearance <- "SDC\_EDIT"
      ProcessValue <- "DB_SDC_GLOBAL_START_COURSE"
      ObjectEnable <- "SDC\_EDIT"
   TextField "Textfeld_9" at 109,351 size 170x31; Text 'track start [mm] / Start Course mm / Track Start [mm]'
   IOField "EA-Feld_12" at 245,350 size 122x32; FormatPattern 99999999
      Appearance <- "SDC\_EDIT"
      ProcessValue <- "DB_SDC_GLOBAL_END_COURSE"
      ObjectEnable <- "SDC\_EDIT"
   TextField "Textfeld_11" at 446,352 size 178x31; Text 'track end [mm] / End Course mm / Track End [mm]'
   TextField "Textfeld_1" at 480,429 size 243x27; Text 'section counter / min Barcode mm / Production zone spacing'
   TextField "Textfeld_2" at 480,469 size 315x27; Text 'EMS No. with vacuum cleaner / min Barcode mm / Accum zone spacing'
   IOField "EA-Feld_1" at 406,424 size 61x32; FormatPattern 9999
      ProcessValue <- "EMS_Production_Spacing"
      Appearance <- "EMS_Production_Spacing"
   IOField "EA-Feld_2" at 406,466 size 61x32; FormatPattern 9999
      ProcessValue <- "EMS_Carrier_Spacing"
      Appearance <- "EMS_Carrier_Spacing"
   TextField "Textfeld_3" at 881,262 size 243x27; Text 'section counter / min Barcode mm / Production zone speed'
   TextField "Textfeld_4" at 881,302 size 315x27; Text 'EMS No. with vacuum cleaner / min Barcode mm / Accum zone speed'
   IOField "EA-Feld_3" at 807,257 size 61x32; FormatPattern 9999
      ProcessValue <- "EMS_Production_Zone_Speed"
      Appearance <- "EMS_Production_Spacing"
   IOField "EA-Feld_4" at 807,299 size 61x32; FormatPattern 99999
      ProcessValue <- "EMS_Accum_Zone_Speed"
      Appearance <- "EMS_Carrier_Spacing"
   TextField "Textfeld_5" at 881,347 size 243x27; Text 'section counter / min Barcode mm / Coarse decel speed'
   TextField "Textfeld_6" at 881,387 size 315x27; Text 'EMS No. with vacuum cleaner / min Barcode mm / Fine decel speed'
   IOField "EA-Feld_5" at 807,342 size 61x32; FormatPattern 9999
      ProcessValue <- "EMS_Coarse_Decel_Speed"
      Appearance <- "EMS_Production_Spacing"
   IOField "EA-Feld_6" at 807,384 size 61x32; FormatPattern 99999
      ProcessValue <- "EMS_Fine_Decel_Speed"
      Appearance <- "EMS_Carrier_Spacing"
   TextField "Textfeld_7" at 881,429 size 243x27; Text 'section counter / min Barcode mm / Coarse position tolerance'
   TextField "Textfeld_8" at 881,469 size 315x27; Text 'EMS No. with vacuum cleaner / min Barcode mm / Fine position tolerance'
   IOField "EA-Feld_7" at 807,424 size 61x32; FormatPattern 9999
      ProcessValue <- "EMS_Coarse_Position_Tolerance"
      Appearance <- "EMS_Production_Spacing"
   IOField "EA-Feld_8" at 807,466 size 61x32; FormatPattern 99999
      ProcessValue <- "EMS_Fine_Posistion_Tolerance"
      Appearance <- "EMS_Carrier_Spacing"
   TextField "Textfeld_10" at 881,511 size 243x27; Text 'section counter / min Barcode mm / Coarse position decel offset'
   TextField "Textfeld_12" at 881,551 size 315x27; Text 'EMS No. with vacuum cleaner / min Barcode mm / Fine position decel offset'
   IOField "EA-Feld_9" at 807,506 size 61x32; FormatPattern 9999
      ProcessValue <- "EMS_Coarse_Position_Decel_Offset"
      Appearance <- "EMS_Production_Spacing"
   IOField "EA-Feld_11" at 807,548 size 61x32; FormatPattern 99999
      ProcessValue <- "EMS_Fine_Position_Decel_Offset"
      Appearance <- "EMS_Carrier_Spacing"
   TextField "Textfeld_13" at 568,143 size 243x27; Text 'section counter / min Barcode mm / Global Parameter'

